// TIA Portal project "management parcare auto" (V17) (continued)
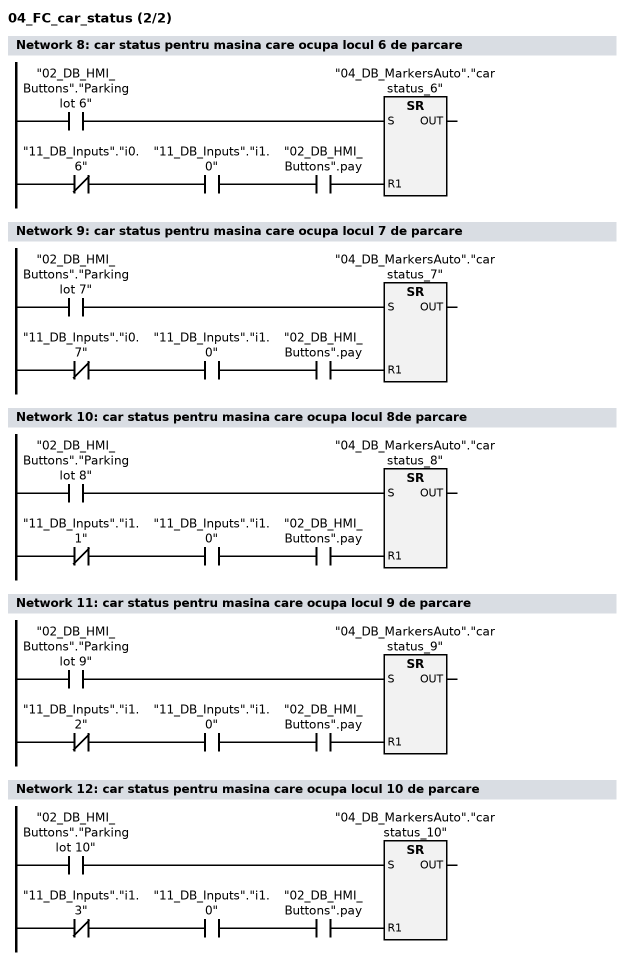
   RUNG wire#powerrail
      Contact( "02_DB_HMI_Buttons"."Parking lot 6" )
      S_SR(operand := "04_DB_MarkersAuto"."car status_6", r1 := wire#w1)
   END_RUNG
   RUNG wire#powerrail
      I_Contact( "11_DB_Inputs"."i0.6" )
      Contact( "11_DB_Inputs"."i1.0" )
      Contact( "02_DB_HMI_Buttons".pay )
   END_RUNG wire#w1
   // the same network as SCL:
   IF "02_DB_HMI_Buttons"."Parking lot 6" THEN
       "04_DB_MarkersAuto"."car status_6" := TRUE;   // SR flip-flop
   END_IF;
   IF NOT "11_DB_Inputs"."i0.6" AND "11_DB_Inputs"."i1.0" AND "02_DB_HMI_Buttons".pay THEN
       "04_DB_MarkersAuto"."car status_6" := FALSE;
   END_IF;
END_REGION

REGION Network 9: car status pentru masina care ocupa locul 7 de parcare
   RUNG wire#powerrail
      Contact( "02_DB_HMI_Buttons"."Parking lot 7" )
      S_SR(operand := "04_DB_MarkersAuto"."car status_7", r1 := wire#w1)
   END_RUNG
   RUNG wire#powerrail
      I_Contact( "11_DB_Inputs"."i0.7" )
      Contact( "11_DB_Inputs"."i1.0" )
      Contact( "02_DB_HMI_Buttons".pay )
   END_RUNG wire#w1
   // the same network as SCL:
   IF "02_DB_HMI_Buttons"."Parking lot 7" THEN
       "04_DB_MarkersAuto"."car status_7" := TRUE;   // SR flip-flop
   END_IF;
   IF NOT "11_DB_Inputs"."i0.7" AND "11_DB_Inputs"."i1.0" AND "02_DB_HMI_Buttons".pay THEN
       "04_DB_MarkersAuto"."car status_7" := FALSE;
   END_IF;
END_REGION

REGION Network 10: car status pentru masina care ocupa locul 8de parcare
   RUNG wire#powerrail
      Contact( "02_DB_HMI_Buttons"."Parking lot 8" )
      S_SR(operand := "04_DB_MarkersAuto"."car status_8", r1 := wire#w1)
   END_RUNG
   RUNG wire#powerrail
      I_Contact( "11_DB_Inputs"."i1.1" )
      Contact( "11_DB_Inputs"."i1.0" )
      Contact( "02_DB_HMI_Buttons".pay )
   END_RUNG wire#w1
   // the same network as SCL:
   IF "02_DB_HMI_Buttons"."Parking lot 8" THEN
       "04_DB_MarkersAuto"."car status_8" := TRUE;   // SR flip-flop
   END_IF;
   IF NOT "11_DB_Inputs"."i1.1" AND "11_DB_Inputs"."i1.0" AND "02_DB_HMI_Buttons".pay THEN
       "04_DB_MarkersAuto"."car status_8" := FALSE;
   END_IF;
END_REGION

REGION Network 11: car status pentru masina care ocupa locul 9 de parcare
   RUNG wire#powerrail
      Contact( "02_DB_HMI_Buttons"."Parking lot 9" )
      S_SR(operand := "04_DB_MarkersAuto"."car status_9", r1 := wire#w1)
   END_RUNG
   RUNG wire#powerrail
      I_Contact( "11_DB_Inputs"."i1.2" )
      Contact( "11_DB_Inputs"."i1.0" )
      Contact( "02_DB_HMI_Buttons".pay )
   END_RUNG wire#w1
   // the same network as SCL:
   IF "02_DB_HMI_Buttons"."Parking lot 9" THEN
       "04_DB_MarkersAuto"."car status_9" := TRUE;   // SR flip-flop
   END_IF;
   IF NOT "11_DB_Inputs"."i1.2" AND "11_DB_Inputs"."i1.0" AND "02_DB_HMI_Buttons".pay THEN
       "04_DB_MarkersAuto"."car status_9" := FALSE;
   END_IF;
END_REGION

REGION Network 12: car status pentru masina care ocupa locul 10 de parcare
   RUNG wire#powerrail
      Contact( "02_DB_HMI_Buttons"."Parking lot 10" )
      S_SR(operand := "04_DB_MarkersAuto"."car status_10", r1 := wire#w1)
   END_RUNG
   RUNG wire#powerrail
      I_Contact( "11_DB_Inputs"."i1.3" )
      Contact( "11_DB_Inputs"."i1.0" )
      Contact( "02_DB_HMI_Buttons".pay )
   END_RUNG wire#w1
   // the same network as SCL:
   IF "02_DB_HMI_Buttons"."Parking lot 10" THEN
       "04_DB_MarkersAuto"."car status_10" := TRUE;   // SR flip-flop
   END_IF;
   IF NOT "11_DB_Inputs"."i1.3" AND "11_DB_Inputs"."i1.0" AND "02_DB_HMI_Buttons".pay THEN
       "04_DB_MarkersAuto"."car status_10" := FALSE;
   END_IF;
END_REGION
END_FUNCTION

FUNCTION "05_FC_Alarms" : Void   // FC5, LAD
{ S7_Optimized_Access := 'TRUE' }
VERSION : 0.1
BEGIN

REGION Network 1: parcare full=> nu are voie sa intre in parcare
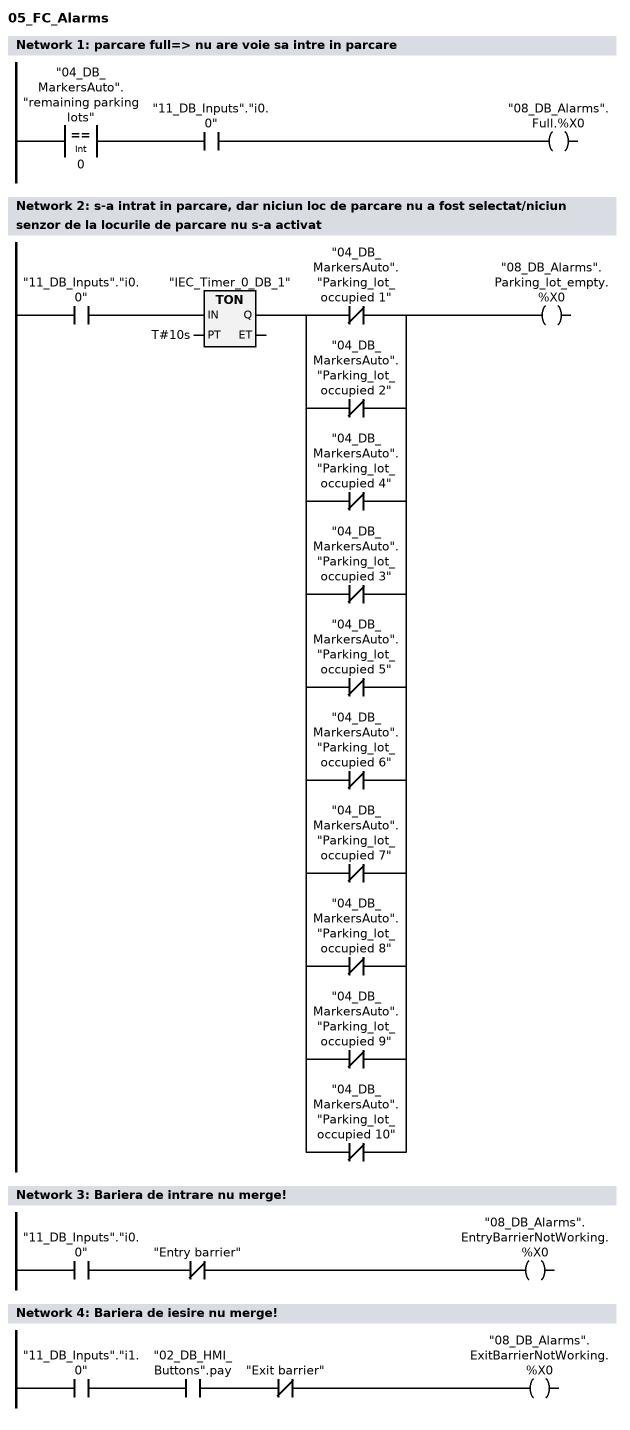
   RUNG wire#powerrail
      { S7_Templates := "SrcType := Int" } EQ_Contact(in1 := "04_DB_MarkersAuto"."remaining parking lots", in2 := 0)
      Contact( "11_DB_Inputs"."i0.0" )
      Coil( "08_DB_Alarms".Full.%X0 )
   END_RUNG
   // the same network as SCL:
   "08_DB_Alarms".Full.%X0 := ("04_DB_MarkersAuto"."remaining parking lots" = 0) AND "11_DB_Inputs"."i0.0";
END_REGION

REGION Network 2: s-a intrat in parcare, dar niciun loc de parcare nu a fost selectat/niciun senzor de la locurile de parcare nu s-a activat
   "IEC_Timer_0_DB_1".TON(IN := "11_DB_Inputs"."i0.0", PT := T#10s);
   "08_DB_Alarms".Parking_lot_empty.%X0 := "IEC_Timer_0_DB_1".Q AND (NOT "04_DB_MarkersAuto"."Parking_lot_occupied 1" OR NOT "04_DB_MarkersAuto"."Parking_lot_occupied 2" OR NOT "04_DB_MarkersAuto"."Parking_lot_occupied 4" OR NOT "04_DB_MarkersAuto"."Parking_lot_occupied 3" OR NOT "04_DB_MarkersAuto"."Parking_lot_occupied 5" OR NOT "04_DB_MarkersAuto"."Parking_lot_occupied 6" OR NOT "04_DB_MarkersAuto"."Parking_lot_occupied 7" OR NOT "04_DB_MarkersAuto"."Parking_lot_occupied 8" OR NOT "04_DB_MarkersAuto"."Parking_lot_occupied 9" OR NOT "04_DB_MarkersAuto"."Parking_lot_occupied 10");
END_REGION

REGION Network 3: Bariera de intrare nu merge!
   RUNG wire#powerrail
      Contact( "11_DB_Inputs"."i0.0" )
      I_Contact( "Entry barrier" )
      Coil( "08_DB_Alarms".EntryBarrierNotWorking.%X0 )
   END_RUNG
   // the same network as SCL:
   "08_DB_Alarms".EntryBarrierNotWorking.%X0 := "11_DB_Inputs"."i0.0" AND NOT "Entry barrier";
END_REGION

REGION Network 4: Bariera de iesire nu merge!
   RUNG wire#powerrail
      Contact( "11_DB_Inputs"."i1.0" )
      Contact( "02_DB_HMI_Buttons".pay )
      I_Contact( "Exit barrier" )
      Coil( "08_DB_Alarms".ExitBarrierNotWorking.%X0 )
   END_RUNG
   // the same network as SCL:
   "08_DB_Alarms".ExitBarrierNotWorking.%X0 := "11_DB_Inputs"."i1.0" AND "02_DB_HMI_Buttons".pay AND NOT "Exit barrier";
END_REGION
END_FUNCTION

FUNCTION "06_FC_Entry_logic" : Void   // FC6, LAD
{ S7_Optimized_Access := 'TRUE' }
VERSION : 0.1
BEGIN

REGION Network 1
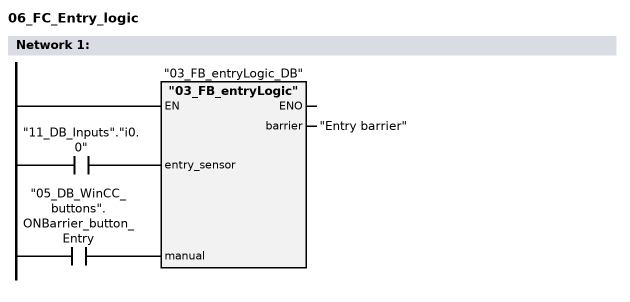
   RUNG wire#powerrail
      "03_FB_entryLogic_DB"(entry_sensor := wire#w1, manual := wire#w2, barrier => "Entry barrier")
   END_RUNG
   RUNG wire#powerrail
      Contact( "11_DB_Inputs"."i0.0" )
   END_RUNG wire#w1
   RUNG wire#powerrail
      Contact( "05_DB_WinCC_buttons".ONBarrier_button_Entry )
   END_RUNG wire#w2
   // the same network as SCL:
   "03_FB_entryLogic_DB"(entry_sensor := "11_DB_Inputs"."i0.0",   // "03_FB_entryLogic"
                         manual := "05_DB_WinCC_buttons".ONBarrier_button_Entry,
                         barrier => "Entry barrier");
END_REGION
END_FUNCTION

FUNCTION "07_FC_VbScript" : Void   // FC7, LAD
{ S7_Optimized_Access := 'TRUE' }
VERSION : 0.1
   VAR_TEMP
      compare : Bool;
   END_VAR
BEGIN

REGION Network 1: tagg folosit ca trigger pentru a rula vbScriptul
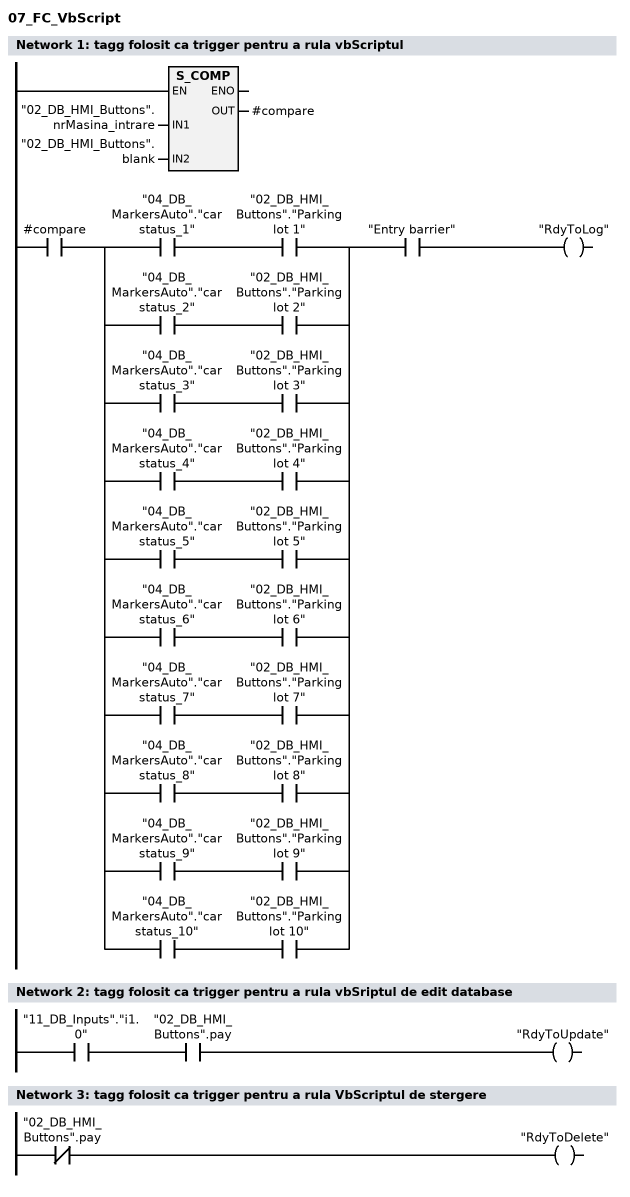
   S_COMP(IN1 := "02_DB_HMI_Buttons".nrMasina_intrare, IN2 := "02_DB_HMI_Buttons".blank, OUT => #compare);
   "RdyToLog" := #compare AND (("04_DB_MarkersAuto"."car status_1" AND "02_DB_HMI_Buttons"."Parking lot 1") OR ("04_DB_MarkersAuto"."car status_2" AND "02_DB_HMI_Buttons"."Parking lot 2") OR ("04_DB_MarkersAuto"."car status_3" AND "02_DB_HMI_Buttons"."Parking lot 3") OR ("04_DB_MarkersAuto"."car status_4" AND "02_DB_HMI_Buttons"."Parking lot 4") OR ("04_DB_MarkersAuto"."car status_5" AND "02_DB_HMI_Buttons"."Parking lot 5") OR ("04_DB_MarkersAuto"."car status_6" AND "02_DB_HMI_Buttons"."Parking lot 6") OR ("04_DB_MarkersAuto"."car status_7" AND "02_DB_HMI_Buttons"."Parking lot 7") OR ("04_DB_MarkersAuto"."car status_8" AND "02_DB_HMI_Buttons"."Parking lot 8") OR ("04_DB_MarkersAuto"."car status_9" AND "02_DB_HMI_Buttons"."Parking lot 9") OR ("04_DB_MarkersAuto"."car status_10" AND "02_DB_HMI_Buttons"."Parking lot 10")) AND "Entry barrier";
END_REGION

REGION Network 2: tagg folosit ca trigger pentru a rula vbSriptul de edit database
   RUNG wire#powerrail
      Contact( "11_DB_Inputs"."i1.0" )
      Contact( "02_DB_HMI_Buttons".pay )
      Coil( "RdyToUpdate" )
   END_RUNG
   // the same network as SCL:
   "RdyToUpdate" := "11_DB_Inputs"."i1.0" AND "02_DB_HMI_Buttons".pay;
END_REGION

REGION Network 3: tagg folosit ca trigger pentru a rula VbScriptul de stergere
   RUNG wire#powerrail
      I_Contact( "02_DB_HMI_Buttons".pay )
      Coil( "RdyToDelete" )
   END_RUNG
   // the same network as SCL:
   "RdyToDelete" := NOT "02_DB_HMI_Buttons".pay;
END_REGION
END_FUNCTION

(* ===== HMI "HMI_RT_1" =====
system functions are stored by id; their names below are inferred from use
connection "HMI_Connection_2": ETHERNET, S7_1500_OMS

HMI tags "Default tag table"
   "04_DB_MarkersAuto_car status_1" : Bool = PLC "04_DB_MarkersAuto"."car status_1" AT %DB1.DBX0.0, 1 s
   "02_DB_HMI_Buttons_nr_masina" : String[254] = PLC "02_DB_HMI_Buttons".nrMasina_intrare AT %DB1.DBX0.0, 1 s
   "RdyToLog" : Bool = PLC RdyToLog AT %M2.0, 100 ms
      on ChangeValue: "Insert_to_database"()
   "Parking lot 1 sensor" : Bool = PLC "11_DB_Inputs"."i0.1" AT %DB1.DBX0.0, 1 s
   "Parking lot 2 sensor" : Bool = PLC "11_DB_Inputs"."i0.2" AT %DB1.DBX0.0, 1 s
   "Parking lot 3 sensor" : Bool = PLC "11_DB_Inputs"."i0.3" AT %DB1.DBX0.0, 1 s
   "Parking lot 4 sensor" : Bool = PLC "11_DB_Inputs"."i0.4" AT %DB1.DBX0.0, 1 s
   "Parking lot 5 sensor" : Bool = PLC "11_DB_Inputs"."i0.5" AT %DB1.DBX0.0, 1 s
   "Parking lot 6 sensor" : Bool = PLC "11_DB_Inputs"."i0.6" AT %DB1.DBX0.0, 1 s
   "Parking lot 7 sensor" : Bool = PLC "11_DB_Inputs"."i0.7" AT %DB1.DBX0.0, 1 s
   "Parking lot 8 sensor" : Bool = PLC "11_DB_Inputs"."i1.1" AT %DB1.DBX0.0, 1 s
   "Parking lot 9 sensor" : Bool = PLC "11_DB_Inputs"."i1.2" AT %DB1.DBX0.0, 1 s
   "Parking lot 10 sensor" : Bool = PLC "11_DB_Inputs"."i1.3" AT %DB1.DBX0.0, 1 s
   "Entry barrier" : Bool = PLC "Entry barrier" AT %Q0.0, 1 s
   "Exit barrier" : Bool = PLC "Exit barrier" AT %Q0.1, 1 s
   "04_DB_MarkersAuto_car status_2" : Bool = PLC "04_DB_MarkersAuto"."car status_2" AT %DB1.DBX0.0, 1 s
   "04_DB_MarkersAuto_car status_3" : Bool = PLC "04_DB_MarkersAuto"."car status_3" AT %DB1.DBX0.0, 1 s
   "04_DB_MarkersAuto_car status_4" : Bool = PLC "04_DB_MarkersAuto"."car status_4" AT %DB1.DBX0.0, 1 s
   "04_DB_MarkersAuto_car status_5" : Bool = PLC "04_DB_MarkersAuto"."car status_5" AT %DB1.DBX0.0, 1 s
   "04_DB_MarkersAuto_car status_6" : Bool = PLC "04_DB_MarkersAuto"."car status_6" AT %DB1.DBX0.0, 1 s
   "04_DB_MarkersAuto_car status_7" : Bool = PLC "04_DB_MarkersAuto"."car status_7" AT %DB1.DBX0.0, 1 s
   "04_DB_MarkersAuto_car status_8" : Bool = PLC "04_DB_MarkersAuto"."car status_8" AT %DB1.DBX0.0, 1 s
   "04_DB_MarkersAuto_car status_9" : Bool = PLC "04_DB_MarkersAuto"."car status_9" AT %DB1.DBX0.0, 1 s
   "04_DB_MarkersAuto_car status_10" : Bool = PLC "04_DB_MarkersAuto"."car status_10" AT %DB1.DBX0.0, 1 s
   "02_DB_HMI_Buttons_pay" : Bool = PLC "02_DB_HMI_Buttons".pay AT %DB1.DBX0.0, 1 s
   "02_DB_HMI_Buttons_nrMasina_iesire" : String[254] = PLC "02_DB_HMI_Buttons".nrMasina_iesire AT %DB1.DBX0.0, 1 s
   "RdyToUpdate" : Bool = PLC RdyToUpdate AT %M6.0, 100 ms
      on ChangeValue: "EditDataRecord"()
   "11_DB_Inputs_i0.0" : Bool = PLC "11_DB_Inputs"."i0.0" AT %DB1.DBX0.0, 1 s
   "11_DB_Inputs_i1.0" : Bool = PLC "11_DB_Inputs"."i1.0" AT %DB1.DBX0.0, 1 s
   "RdyToDelete" : Bool = PLC RdyToDelete AT %M6.1, 100 ms
      on ChangeValue: "Delete_from_database"()
   "Numar_masini_ziuaX" : Int, internal
   "filtrare_dupa_data" : WString[254], internal
   "Interval1_date" : WString[254], internal
   "Interval2_date" : WString[254], internal
   "nr_masini_interval" : Int, internal
   "nr_total_masini" : Int, internal
   "Verficare_rulareScriptInsr" : Bool = PLC "05_DB_WinCC_buttons".ResetNumber AT %DB1.DBX0.0, 1 s
   "EntrButton_ON" : Bool = PLC "05_DB_WinCC_buttons".ONBarrier_button_Entry AT %DB1.DBX0.0, 1 s
   "ExitButton_ON" : Bool = PLC "05_DB_WinCC_buttons".ONBarrier_button_Exit AT %DB1.DBX0.0, 1 s

HMI tags "Read_temp"
   "CarStatus1" : Int, internal
   "CarStatus2" : Int, internal
   "CarStatus3" : Int, internal
   "CarStatus4" : Int, internal
   "CarStatus5" : Int, internal
   "CarStatus7" : Int, internal
   "CarStatus8" : Int, internal
   "CarStatus9" : Int, internal
   "CarStatus10" : Int, internal
   "OraIntrare1" : DateTime, internal
   "OraIntrare2" : DateTime, internal
   "OraIntrare3" : DateTime, internal
   "OraIntrare4" : DateTime, internal
   "OraIntrare5" : DateTime, internal
   "OraIntrare6" : DateTime, internal
   "OraIntrare7" : DateTime, internal
   "OraIntrare8" : DateTime, internal
   "OraIntrare9" : DateTime, internal
   "OraIntrare10" : DateTime, internal
   "CarStatus6" : Int, internal
   "DataIntrare1" : DateTime, internal
   "DataIntrare2" : DateTime, internal
   "DataIntrare3" : DateTime, internal
   "DataIntrare4" : DateTime, internal
   "DataIntrare5" : DateTime, internal
   "DataIntrare6" : DateTime, internal
   "DataIntrare7" : DateTime, internal
   "DataIntrare8" : DateTime, internal
   "DataIntrare9" : DateTime, internal
   "DataIntrare10" : DateTime, internal
   "OraIesire1" : DateTime, internal
   "OraIesire2" : DateTime, internal
   "OraIesire3" : DateTime, internal
   "OraIesire4" : DateTime, internal
   "OraIesire5" : DateTime, internal
   "OraIesire6" : DateTime, internal
   "OraIesire7" : DateTime, internal
   "OraIesire8" : DateTime, internal
   "OraIesire9" : DateTime, internal
   "OraIesire10" : DateTime, internal
   "DataIesire1" : DateTime, internal
   "DataIesire2" : DateTime, internal
   "DataIesire3" : DateTime, internal
   "DataIesire4" : DateTime, internal
   "DataIesire5" : DateTime, internal
   "DataIesire6" : DateTime, internal
   "DataIesire7" : DateTime, internal
   "DataIesire8" : DateTime, internal
   "DataIesire9" : DateTime, internal
   "DataIesire10" : DateTime, internal
   "NrMasina1" : WString[254], internal
   "NrMasina2" : WString[254], internal
   "NrMasina3" : WString[254], internal
   "NrMasina4" : WString[254], internal
   "NrMasina5" : WString[254], internal
   "NrMasina6" : WString[254], internal
   "NrMasina7" : WString[254], internal
   "NrMasina8" : WString[254], internal
   "NrMasina9" : WString[254], internal
   "NrMasina10" : WString[254], internal

HMI tags "Read_perm"
   "CarNumber1" : WString[254], internal
   "CarNumber2" : WString[254], internal
   "CarNumber3" : WString[254], internal
   "CarNumber4" : WString[254], internal
   "CarNumber5" : WString[254], internal
   "CarNumber6" : WString[254], internal
   "CarNumber7" : WString[254], internal
   "CarNumber8" : WString[254], internal
   "CarNumber9" : WString[254], internal
   "CarNumber10" : WString[254], internal
   "Status1" : Int, internal
   "Status2" : Int, internal
   "Status3" : Int, internal
   "Status4" : Int, internal
   "Status5" : Int, internal
   "Status6" : Int, internal
   "Status7" : Int, internal
   "Status8" : Int, internal
   "Status9" : Int, internal
   "Status10" : Int, internal
   "EntryTime1" : DateTime, internal
   "EntryTime2" : DateTime, internal
   "EntryTime3" : DateTime, internal
   "EntryTime4" : DateTime, internal
   "EntryTime5" : DateTime, internal
   "EntryTime6" : DateTime, internal
   "EntryTime7" : DateTime, internal
   "EntryTime8" : DateTime, internal
   "EntryTime9" : DateTime, internal
   "EntryTime10" : DateTime, internal
   "EntryDate1" : DateTime, internal
   "EntryDate2" : DateTime, internal
   "EntryDate3" : DateTime, internal
   "EntryDate4" : DateTime, internal
   "EntryDate5" : DateTime, internal
   "EntryDate6" : DateTime, internal
   "EntryDate7" : DateTime, internal
   "EntryDate8" : DateTime, internal
   "EntryDate9" : DateTime, internal
   "EntryDate10" : DateTime, internal
   "ExitTime1" : DateTime, internal
   "ExitTime2" : DateTime, internal
   "ExitTime3" : DateTime, internal
   "ExitTime4" : DateTime, internal
   "ExitTime5" : DateTime, internal
   "ExitTime6" : DateTime, internal
   "ExitTime7" : DateTime, internal
   "ExitTime8" : DateTime, internal
   "ExitTime9" : DateTime, internal
   "ExitTime10" : DateTime, internal
   "ExitDate1" : DateTime, internal
   "ExitDate2" : DateTime, internal
   "ExitDate3" : DateTime, internal
   "ExitDate4" : DateTime, internal
   "ExitDate5" : DateTime, internal
   "ExitDate6" : DateTime, internal
   "ExitDate7" : DateTime, internal
   "ExitDate8" : DateTime, internal
   "ExitDate9" : DateTime, internal
   "ExitDate10" : DateTime, internal

HMI tags "Alarms"
   "Alarma_full" : Word = PLC "08_DB_Alarms".Full AT %DB1.DBW0, 1 s
   "Alarma_loc neselectat" : Word = PLC "08_DB_Alarms".Parking_lot_empty AT %DB1.DBW0, 1 s
   "Alarma_barieraIntr_nu" : Word = PLC "08_DB_Alarms".EntryBarrierNotWorking AT %DB1.DBW0, 1 s
   "Alarma_barieraIesire_nu" : Word = PLC "08_DB_Alarms".ExitBarrierNotWorking AT %DB1.DBW0, 1 s

discrete alarms
   1: 'The parking lot is at maximum capacity. You have nowhere to park!', class Warnings, trigger "Alarma_full" bit 0
   2: 'No parking space has been selected. Please select a free parking spot! / Niciun loc de parcare nu a fost selectat. Te rugam sa selectezi un loc liber!', class Warnings, trigger "Alarma_loc neselectat" bit 0
   3: 'The entry barrier does not work! Call the operator!', class Errors, trigger "Alarma_barieraIntr_nu" bit 0
   4: 'The exit barrier does not work! Call the operator!', class Errors, trigger "Alarma_barieraIesire_nu" bit 0

screen "Alarms" 1920x1080
   Button "Button_1" at 1748,4 size 170x79; TextOff 'Exit / Iesire'
      on Press: StopRuntime(0)
   TextField "Text field_1" at 478,90 size 773x166; Text 'Alarms'
   GraphicView "Graphic view_2" at 28,12 size 394x64; Picture "Siemens_AG_logo.svg"
   Button "Button_2" at 9,972 size 194x96; TextOff 'Home / Ecran principal'
      on Press: ActivateScreen("Home", 0)
   AlarmView "Alarm view_1" at 100,217 size 1726x718
   Button "Button_3" at 208,973 size 194x96; TextOff 'Alarms'
      on Press: ActivateScreen("Alarms", 0)
   Button "Button_8" at 408,973 size 194x96; TextOff 'Parking history'
      on Press: ActivateScreen("Parking history", 0)
   Button "Button_4" at 608,973 size 194x96; TextOff 'Statistics'
      on Press: ActivateScreen("Statistics", 0)

screen "Home" 1920x1080
   Button "Button_1" at 1748,4 size 170x79; TextOff 'Exit / Iesire'
      on Press: StopRuntime(0)
   TextField "Text field_1" at 469,95 size 869x186; Text 'Parking car'
   TextField "Text field_2" at 302,224 size 437x47; Text 'SENSOR STATUS / Status Senzori'
   TextField "Text field_3" at 142,366 size 93x104; Text 'Entry sensor'
   TextField "Text field_4" at 285,364 size 93x104; Text 'Exit sensor'
   TextField "Text field_5" at 469,265 size 93x104; Text 'No. 1 sensor'
   TextField "Text field_6" at 469,332 size 93x104; Text 'No. 2 sensor'
   TextField "Text field_7" at 473,422 size 19x29; Text 'Text'
   TextField "Text field_8" at 469,406 size 93x104; Text 'No. 3 sensor'
   TextField "Text field_9" at 467,473 size 93x104; Text 'No. 4 sensor'
   TextField "Text field_10" at 467,543 size 93x104; Text 'No. 5 sensor'
   TextField "Text field_11" at 664,262 size 93x104; Text 'No. 6 sensor'
   TextField "Text field_12" at 664,330 size 93x104; Text 'No. 7 sensor'
   TextField "Text field_13" at 662,401 size 93x104; Text 'No. 8 sensor'
   TextField "Text field_14" at 662,472 size 93x104; Text 'No. 9 sensor'
   TextField "Text field_15" at 664,538 size 93x104; Text 'No. 10 sensor'
   Ellipse "Ellipse_1" at 562,293 size 52x50
      Appearance <- "Parking lot 1 sensor"
   Ellipse "Ellipse_2" at 561,361 size 52x50
      Appearance <- "Parking lot 2 sensor"
   Ellipse "Ellipse_3" at 560,431 size 52x50
      Appearance <- "Parking lot 3 sensor"
   Ellipse "Ellipse_4" at 559,501 size 52x50
      Appearance <- "Parking lot 4 sensor"
   Ellipse "Ellipse_5" at 558,570 size 52x50
      Appearance <- "Parking lot 5 sensor"
   Ellipse "Ellipse_6" at 752,290 size 52x50
      Appearance <- "Parking lot 6 sensor"
   Ellipse "Ellipse_7" at 752,360 size 52x50
      Appearance <- "Parking lot 7 sensor"
   Ellipse "Ellipse_8" at 752,430 size 52x50
      Appearance <- "Parking lot 8 sensor"
   Ellipse "Ellipse_9" at 752,499 size 52x50
      Appearance <- "Parking lot 9 sensor"
   Ellipse "Ellipse_10" at 752,568 size 52x50
      Appearance <- "Parking lot 10 sensor"
   Ellipse "Ellipse_11" at 138,452 size 69x67
      Appearance <- "11_DB_Inputs_i0.0"
   Ellipse "Ellipse_12" at 292,451 size 69x67
      Appearance <- "11_DB_Inputs_i1.0"
   GraphicView "Graphic view_2" at 28,12 size 394x64; Picture "Siemens_AG_logo.svg"
   Button "Button_2" at 208,973 size 194x96; TextOff 'Alarms'
      on Press: ActivateScreen("Alarms", 0)
   TextField "Text field_16" at 1162,185 size 581x219; Text 'LIVE BARRIERS'
   GraphicView "Graphic view_3" at 1525,515 size 56x80; Picture "pngegg"
   GraphicView "Graphic view_4" at 1186,351 size 56x80; Picture "pngegg"
   GraphicView "Graphic view_5" at 1170,283 size 93x85; Picture "exit"
   GraphicView "Graphic view_6" at 1675,500 size 101x105; Picture "parking"
   TextField "Text field_17" at 761,660 size 437x47; Text 'REMOTE CONTROL / Control Operator'
   TextField "Text field_18" at 585,713 size 453x103; Text 'Entry barrier:'
   TextField "Text field_19" at 586,778 size 341x103; Text 'Exit barrier:'
   Button "Button_8" at 408,973 size 194x96; TextOff 'Parking history'
      on Press: ActivateScreen("Parking history", 0)
   Button "Button_9" at 9,972 size 194x96; TextOff 'Home / Ecran principal'
      on Press: ActivateScreen("Home", 0)
   Line "Line_2" at 1541,520 size 140x0
      Visibility <- "Entry barrier"
   Line "Line_3" at 1202,356 size 140x0
      Visibility <- "Exit barrier"
   Button "Button_3" at 608,973 size 194x96; TextOff 'Statistics'
      on Press: ActivateScreen("Statistics", 0)
   Button "Button_4" at 970,737 size 134x52; TextOff 'ON'
      on Press: SetBit("EntrButton_ON")
      Appearance <- "Entry barrier"
   Button "Button_5" at 970,805 size 134x52; TextOn 'ON'; TextOff 'ON'
      on Press: SetBit("ExitButton_ON")
      Appearance <- "Exit barrier"
   Button "Button_6" at 1128,737 size 134x52; TextOn 'ON'; TextOff 'OFF'
      on Press: ResetBit("EntrButton_ON")
      Appearance <- "Entry barrier"
   Button "Button_7" at 1128,805 size 134x52; TextOn 'ON'; TextOff 'OFF'
      on Press: ResetBit("ExitButton_ON")
      Appearance <- "Exit barrier"
   TextField "Text field_20" at 84,317 size 325x73; Text 'Sensor barriers'
   TextField "Text field_21" at 302,224 size 437x47; Text 'SENSOR STATUS / Status Senzori'
   TextField "Text field_22" at 401,239 size 73x405; Text 'Sensor parking lots'

screen "Parking history" 1920x1080
   on GenerateScreen: "Read_fromTEMP"(); "Read_fromPerm"()
   TextField "Text field_2" at 159,243 size 143x50; Text 'Car status Status Senzori'
   GraphicView "Graphic view_2" at 28,12 size 394x64; Picture "Siemens_AG_logo.svg"
   Button "Button_1" at 1748,4 size 170x79; TextOff 'Exit / Iesire'
      on Press: StopRuntime(0)
   Button "Button_2" at 9,972 size 194x96; TextOff 'Home / Ecran principal'
      on Press: ActivateScreen("Home", 0)
   Button "Button_3" at 208,973 size 194x96; TextOff 'Alarms'
      on Press: ActivateScreen("Alarms", 0)
   Button "Button_8" at 408,973 size 194x96; TextOff 'Parking history'
      on Press: ActivateScreen("Parking history", 0)
   IOField "I/O field_1" at 21,294 size 146x54; FormatPattern ????????
      ProcessValue <- "NrMasina1"
   IOField "I/O field_2" at 163,294 size 109x54; FormatPattern 9
      ProcessValue <- "CarStatus1"
   IOField "I/O field_3" at 268,294 size 172x54; FormatPattern 9999999999999999999999999999999999999999
      ProcessValue <- "OraIntrare1"
   TextField "Text field_1" at 49,221 size 165x119; Text 'Car number'
   IOField "I/O field_5" at 435,294 size 172x54; FormatPattern 9999999999999999999999999999999999999999
      ProcessValue <- "DataIntrare1"
   TextField "Text field_7" at 383,208 size 325x96; Text 'Entry date'
   IOField "I/O field_7" at 21,343 size 149x54; FormatPattern ????????
      ProcessValue <- "NrMasina2"
   IOField "I/O field_8" at 163,343 size 109x54; FormatPattern 9
      ProcessValue <- "CarStatus2"
   IOField "I/O field_9" at 268,343 size 172x54; FormatPattern 9999999999999999999999999999999999999999
      ProcessValue <- "OraIntrare2"
   IOField "I/O field_10" at 435,343 size 172x54; FormatPattern 9999999999999999999999999999999999999999
      ProcessValue <- "DataIntrare2"
   IOField "I/O field_29" at 268,392 size 172x54; FormatPattern 9999999999999999999999999999999999999999
      ProcessValue <- "OraIntrare3"
   IOField "I/O field_30" at 268,441 size 172x54; FormatPattern 9999999999999999999999999999999999999999
      ProcessValue <- "OraIntrare4"
   IOField "I/O field_31" at 268,490 size 172x54; FormatPattern 9999999999999999999999999999999999999999
      ProcessValue <- "OraIntrare5"
   IOField "I/O field_32" at 268,539 size 172x54; FormatPattern 9999999999999999999999999999999999999999
      ProcessValue <- "OraIntrare6"
   IOField "I/O field_33" at 268,588 size 172x54; FormatPattern 9999999999999999999999999999999999999999
      ProcessValue <- "OraIntrare7"
   IOField "I/O field_34" at 268,637 size 172x54; FormatPattern ????
      ProcessValue <- "OraIntrare8"
   IOField "I/O field_35" at 268,686 size 172x54; FormatPattern 9999999999999999999999999999999999999999
      ProcessValue <- "OraIntrare9"
   IOField "I/O field_36" at 268,735 size 172x54; FormatPattern 9999999999999999999999999999999999999999
      ProcessValue <- "OraIntrare10"
   IOField "I/O field_37" at 435,392 size 172x54; FormatPattern 9999999999999999999999999999999999999999
      ProcessValue <- "DataIntrare3"
   IOField "I/O field_38" at 435,441 size 172x54; FormatPattern 9999999999999999999999999999999999999999
      ProcessValue <- "DataIntrare4"
   IOField "I/O field_39" at 435,490 size 172x54; FormatPattern 9999999999999999999999999999999999999999
      ProcessValue <- "DataIntrare5"
   IOField "I/O field_40" at 435,539 size 172x54; FormatPattern 9999999999999999999999999999999999999999
      ProcessValue <- "DataIntrare6"
   IOField "I/O field_41" at 435,588 size 172x54; FormatPattern 9999999999999999999999999999999999999999
      ProcessValue <- "DataIntrare7"
   IOField "I/O field_42" at 435,637 size 172x54; FormatPattern 9999999999999999999999999999999999999999
      ProcessValue <- "DataIntrare8"
   IOField "I/O field_43" at 435,686 size 172x54; FormatPattern 9999999999999999999999999999999999999999
      ProcessValue <- "DataIntrare9"
   IOField "I/O field_44" at 435,735 size 172x54; FormatPattern 9999999999999999999999999999999999999999
      ProcessValue <- "DataIntrare10"
   IOField "I/O field_13" at 21,391 size 149x54; FormatPattern ????????
      ProcessValue <- "NrMasina3"
   IOField "I/O field_14" at 21,439 size 149x54; FormatPattern ????????
      ProcessValue <- "NrMasina4"
   IOField "I/O field_15" at 21,489 size 149x54; FormatPattern ????????
      ProcessValue <- "NrMasina5"
   IOField "I/O field_16" at 21,539 size 149x54; FormatPattern ????????
      ProcessValue <- "NrMasina6"
   IOField "I/O field_17" at 21,588 size 149x54; FormatPattern ????????
      ProcessValue <- "NrMasina7"
   IOField "I/O field_18" at 21,637 size 149x54; FormatPattern ????????
      ProcessValue <- "NrMasina8"
   IOField "I/O field_19" at 21,686 size 149x54; FormatPattern ????????
      ProcessValue <- "NrMasina9"
   IOField "I/O field_20" at 21,735 size 149x54; FormatPattern ????????
      ProcessValue <- "NrMasina10"
   IOField "I/O field_22" at 163,391 size 109x54; FormatPattern 9
      ProcessValue <- "CarStatus3"
   IOField "I/O field_23" at 163,439 size 109x54; FormatPattern 9
      ProcessValue <- "CarStatus4"
   IOField "I/O field_24" at 163,489 size 109x54; FormatPattern 9
      ProcessValue <- "CarStatus5"
   IOField "I/O field_25" at 163,539 size 109x54; FormatPattern 9
      ProcessValue <- "CarStatus6"
   IOField "I/O field_26" at 163,588 size 109x54; FormatPattern 9
      ProcessValue <- "CarStatus7"
   IOField "I/O field_27" at 163,637 size 109x54; FormatPattern 9
      ProcessValue <- "CarStatus8"
   IOField "I/O field_28" at 163,686 size 109x54; FormatPattern 9
      ProcessValue <- "CarStatus9"
   IOField "I/O field_61" at 163,736 size 109x54; FormatPattern 9
      ProcessValue <- "CarStatus10"
   TextField "Text field_9" at 1177,206 size 325x96; Text 'Entry time'
   TextField "Text field_10" at 1355,206 size 325x96; Text 'Entry date'
   TextField "Text field_13" at 1523,207 size 325x96; Text 'Exit time'
   TextField "Text field_5" at 229,210 size 325x96; Text 'Entry time'
   IOField "I/O field_21" at 973,295 size 137x54; FormatPattern ????????
      ProcessValue <- "CarNumber1"
   IOField "I/O field_63" at 1105,295 size 126x54; FormatPattern 9
      ProcessValue <- "Status1"
   IOField "I/O field_64" at 1227,295 size 177x54; FormatPattern 9999999999999999999999999999999999999999
      ProcessValue <- "EntryTime1"
   IOField "I/O field_65" at 1400,295 size 165x54; FormatPattern 9999999999999999999999999999999999999999
      ProcessValue <- "EntryDate1"
   IOField "I/O field_66" at 1562,295 size 164x54; FormatPattern 9999999999999999999999999999999999999999
      ProcessValue <- "ExitTime1"
   IOField "I/O field_62" at 1723,295 size 163x54; FormatPattern 9999999999999999999999999999999999999999
      ProcessValue <- "ExitDate1"
   TextField "Text field_3" at 1049,218 size 165x96; Text 'Car status'
   TextField "Text field_11" at 1669,208 size 245x96; Text 'Exit date'
   Button "Button_4" at 608,973 size 194x96; TextOff 'Statistics'
      on Press: ActivateScreen("Statistics", 0)
   IOField "I/O field_67" at 973,345 size 137x54; FormatPattern ????????
      ProcessValue <- "CarNumber2"
   IOField "I/O field_68" at 973,395 size 137x54; FormatPattern ????????
      ProcessValue <- "CarNumber3"
   IOField "I/O field_69" at 973,445 size 137x54; FormatPattern ????????
      ProcessValue <- "CarNumber4"
   IOField "I/O field_70" at 973,495 size 137x54; FormatPattern ????????
      ProcessValue <- "CarNumber5"
   IOField "I/O field_71" at 973,545 size 137x54; FormatPattern ????????
      ProcessValue <- "CarNumber6"
   IOField "I/O field_72" at 973,595 size 137x54; FormatPattern ????????
      ProcessValue <- "CarNumber7"
   IOField "I/O field_73" at 973,645 size 137x54; FormatPattern ????????
      ProcessValue <- "CarNumber8"
   IOField "I/O field_74" at 973,695 size 137x54; FormatPattern ????????
      ProcessValue <- "CarNumber9"
   IOField "I/O field_75" at 973,745 size 137x54; FormatPattern ????????
      ProcessValue <- "CarNumber10"
   IOField "I/O field_76" at 1105,345 size 126x54; FormatPattern 9